(* Logix 5000 project; controller PLC_MCC1300_75F1 vendor 1 type 14 code 166 rev 32.11; software revision 32.04; part 31 of 83 *)
(* tags used below, declared in another part *)
   B70 : DINT[13];
   BENCH_MASTERUP : ALIAS FOR I[73].6;
   C5 : COUNTER[51];
   I : INT[128];   // Local Input Updates Input Slot 2
   KD_N_MOVIN : ALIAS FOR N14[256].0;
   KD_N_MOVOUT : ALIAS FOR N14[257].0;
   KD_S_MOVIN : ALIAS FOR N14[256].1;
   KD_S_MOVOUT : ALIAS FOR N14[257].1;
   KK_N_MOVDN : ALIAS FOR N14[253].0;
   KK_N_MOVIN : ALIAS FOR N14[254].0;
   KK_N_MOVOUT : ALIAS FOR N14[255].0;
   KK_N_MOVUP : ALIAS FOR N14[252].0;
   KK_S_MOVDN : ALIAS FOR N14[253].1;
   KK_S_MOVIN : ALIAS FOR N14[254].1;
   KK_S_MOVOUT : ALIAS FOR N14[255].1;
   KK_S_MOVUP : ALIAS FOR N14[252].1;
   KNRL_N_AUTO : ALIAS FOR N14[250].0;
   KNRL_N_MANL : ALIAS FOR N14[251].0;
   KNRL_S_AUTO : ALIAS FOR N14[250].1;
   KNRL_S_MANL : ALIAS FOR N14[251].1;
   N11 : DINT[500];
   N12 : DINT[500];
   N14 : DINT[500];
   N214_1 : ALIAS FOR N214[1];
   N26 : DINT[150];
   O : INT[128];
   T4 : TIMER[51];
   TD1_N_MOVIN : ALIAS FOR N14[256].2;
   TD1_N_MOVOUT : ALIAS FOR N14[257].2;
   TD1_S_MOVIN : ALIAS FOR N14[256].3;
   TD1_S_MOVOUT : ALIAS FOR N14[257].3;
   TD2_N_MOVIN : ALIAS FOR N14[256].4;
   TD2_N_MOVOUT : ALIAS FOR N14[257].4;
   TK1_N_MOVDN : ALIAS FOR N14[253].2;
   TK1_N_MOVIN : ALIAS FOR N14[254].2;
   TK1_N_MOVOUT : ALIAS FOR N14[255].2;
   TK1_N_MOVUP : ALIAS FOR N14[252].2;
   TK1_S_MOVDN : ALIAS FOR N14[253].3;
   TK1_S_MOVIN : ALIAS FOR N14[254].3;
   TK1_S_MOVOUT : ALIAS FOR N14[255].3;
   TK1_S_MOVUP : ALIAS FOR N14[252].3;
   TK2_N_MOVDN : ALIAS FOR N14[253].4;
   TK2_N_MOVIN : ALIAS FOR N14[254].4;
   TK2_N_MOVOUT : ALIAS FOR N14[255].4;
   TK2_N_MOVUP : ALIAS FOR N14[252].4;
   TK2_S_MOVDN : ALIAS FOR N14[253].5;
   TK2_S_MOVIN : ALIAS FOR N14[254].5;
   TK2_S_MOVOUT : ALIAS FOR N14[255].5;
   TK2_S_MOVUP : ALIAS FOR N14[252].5;
   TMP_d : DINT;
   TZ1_N_AUTO : ALIAS FOR N14[250].2;
   TZ1_N_MANL : ALIAS FOR N14[251].2;
   TZ1_S_AUTO : ALIAS FOR N14[250].3;
   TZ1_S_MANL : ALIAS FOR N14[251].3;
   TZ2_N_AUTO : ALIAS FOR N14[250].4;
   TZ2_N_MANL : ALIAS FOR N14[251].4;
   TZ2_S_AUTO : ALIAS FOR N14[250].5;
   TZ2_S_MANL : ALIAS FOR N14[251].5;
   VIS_OUTPT_OFF : ALIAS FOR N27[60].2;
   VIS_SYS_STOPPED : ALIAS FOR N27[60].1;
(* MainProgram, continued *)

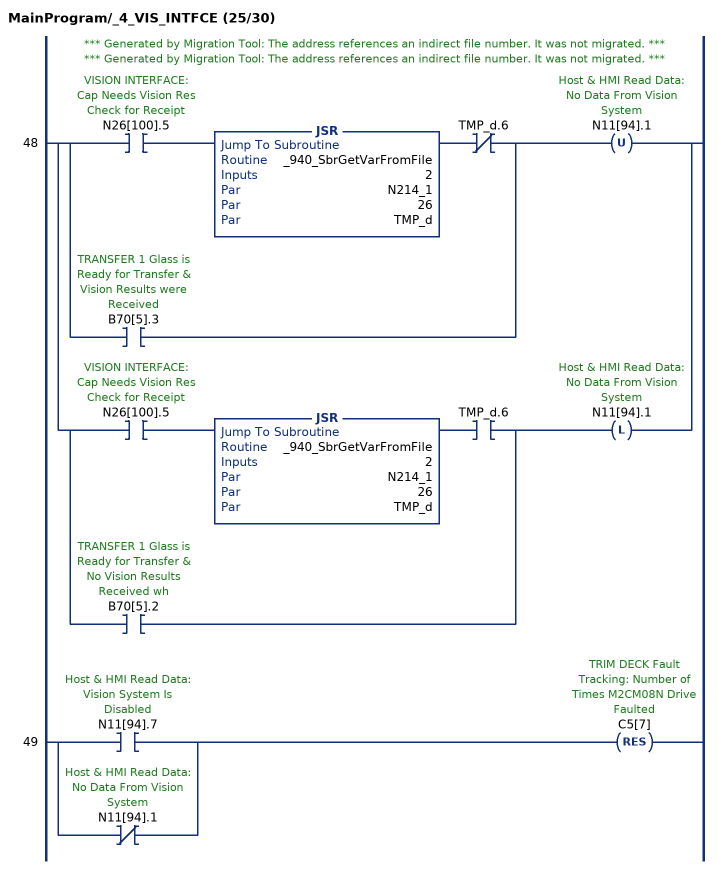
   [picture p426: MainProgram/_4_VIS_INTFCE rungs 48-49]
   // *** Generated by Migration Tool: The address references an indirect file number. It was not migrated. ***
   // *** Generated by Migration Tool: The address references an indirect file number. It was not migrated. ***
   48: [[XIC(N26[100].5) JSR(_940_SbrGetVarFromFile,2,N214_1,26,TMP_d) XIO(TMP_d.6) ,XIC(B70[5].3) ] OTU(N11[94].1) ,[XIC(N26[100].5) JSR(_940_SbrGetVarFromFile,2,N214_1,26,TMP_d) XIC(TMP_d.6) ,XIC(B70[5].2) ] OTL(N11[94].1) ];
   49: [XIC(N11[94].7) ,XIO(N11[94].1) ]RES(C5[7]);
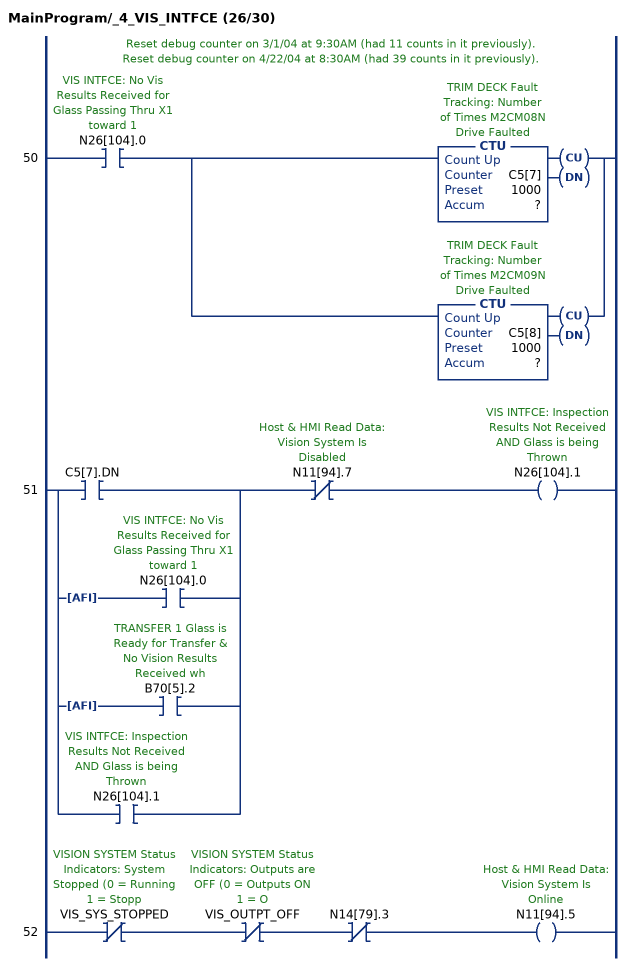
   // Reset debug counter on 3/1/04 at 9:30AM (had 11 counts in it previously).
   // Reset debug counter on 4/22/04 at 8:30AM (had 39 counts in it previously).
   50: XIC(N26[104].0)[CTU(C5[7],?,?) ,CTU(C5[8],?,?) ];
   51: [XIC(C5[7].DN) ,AFI() XIC(N26[104].0) ,AFI() XIC(B70[5].2) ,XIC(N26[104].1) ]XIO(N11[94].7)OTE(N26[104].1);
   52: XIO(VIS_SYS_STOPPED)XIO(VIS_OUTPT_OFF)XIO(N14[79].3)OTE(N11[94].5);
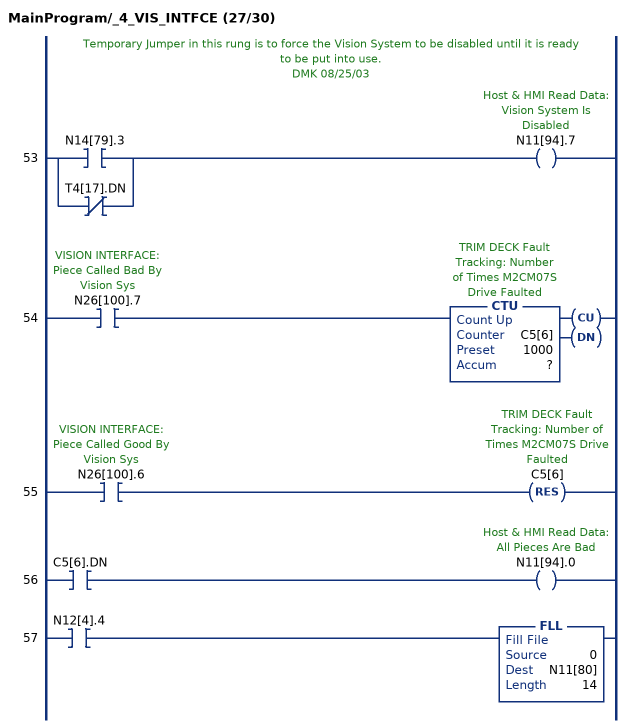
   // Temporary Jumper in this rung is to force the Vision System to be disabled until it is ready to be put into use.
   // DMK 08/25/03
   53: [XIC(N14[79].3) ,XIO(T4[17].DN) ]OTE(N11[94].7);
   54: XIC(N26[100].7)CTU(C5[6],?,?);
   55: XIC(N26[100].6)RES(C5[6]);
   56: XIC(C5[6].DN)OTE(N11[94].0);
   57: XIC(N12[4].4)FLL(0,N11[80],14);
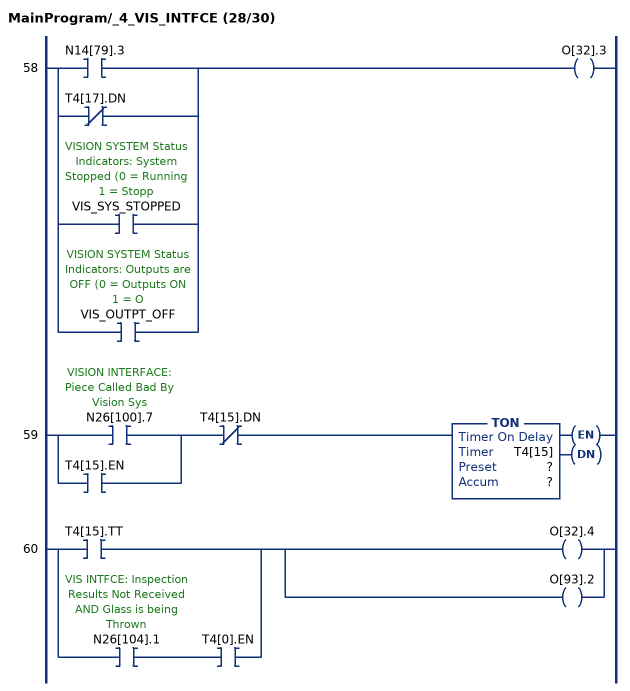
   58: [XIC(N14[79].3) ,XIO(T4[17].DN) ,XIC(VIS_SYS_STOPPED) ,XIC(VIS_OUTPT_OFF) ]OTE(O[32].3);
   59: [XIC(N26[100].7) ,XIC(T4[15].EN) ]XIO(T4[15].DN)TON(T4[15],?,?);
   60: [XIC(T4[15].TT) ,XIC(N26[104].1) XIC(T4[0].EN) ][OTE(O[32].4) ,OTE(O[93].2) ];
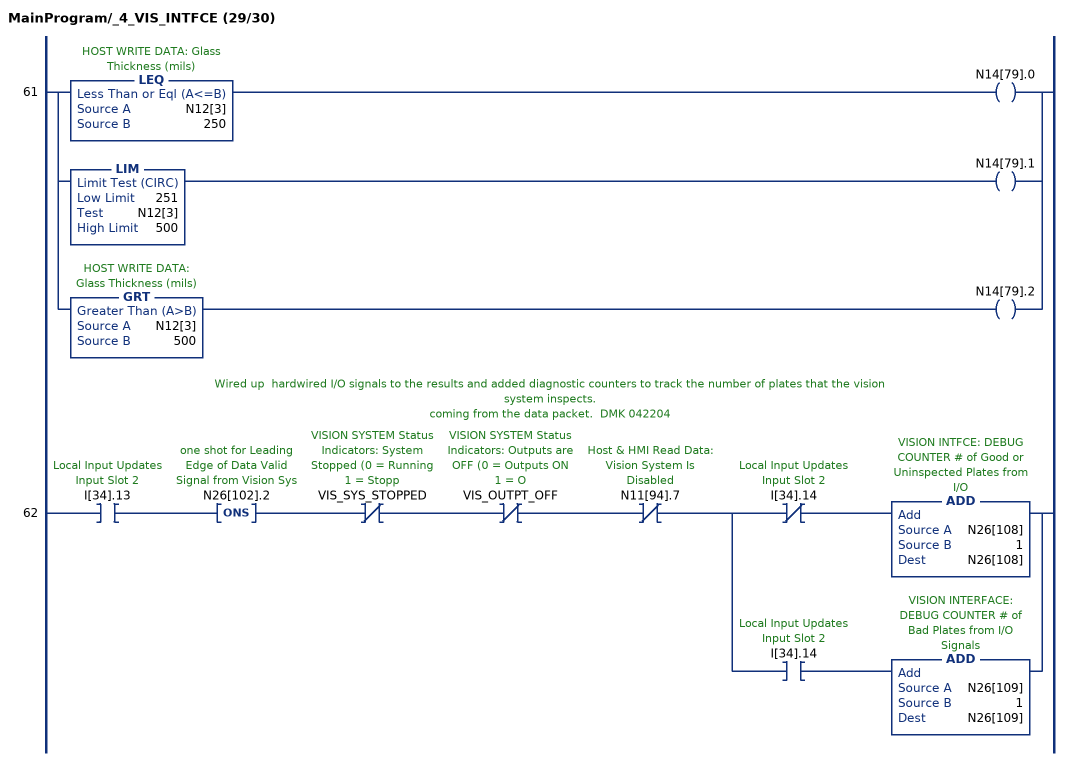
   61: [LEQ(N12[3],250) OTE(N14[79].0) ,LIM(251,N12[3],500) OTE(N14[79].1) ,GRT(N12[3],500) OTE(N14[79].2) ];
   // Wired up  hardwired I/O signals to the results and added diagnostic counters to track the number of plates that the vision
   // system inspects.
   // coming from the data packet.  DMK 042204
   62: XIC(I[34].13)ONS(N26[102].2)XIO(VIS_SYS_STOPPED)XIO(VIS_OUTPT_OFF)XIO(N11[94].7)[XIO(I[34].14) ADD(N26[108],1,N26[108]) ,XIC(I[34].14) ADD(N26[109],1,N26[109]) ];
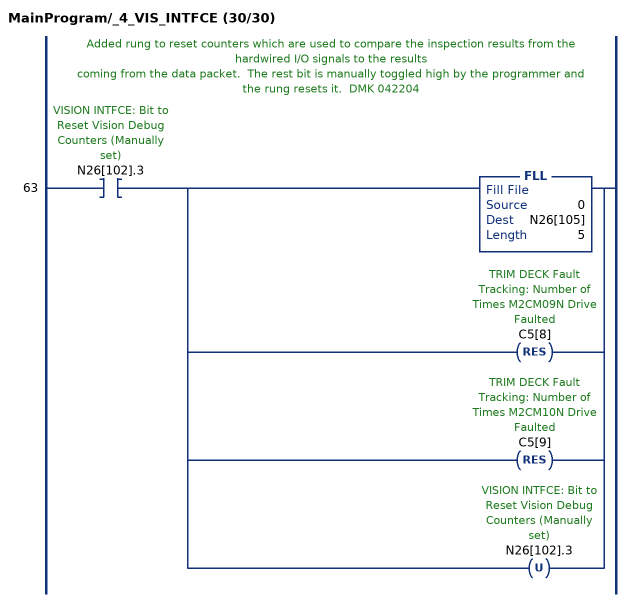
   // Added rung to reset counters which are used to compare the inspection results from the hardwired I/O signals to the results
   // coming from the data packet.  The rest bit is manually toggled high by the programmer and the rung resets it.  DMK 042204
   63: XIC(N26[102].3)[FLL(0,N26[105],5) ,RES(C5[8]) ,RES(C5[9]) ,OTU(N26[102].3) ];
END_ROUTINE

ROUTINE _70_LADDER   (* ladder *)
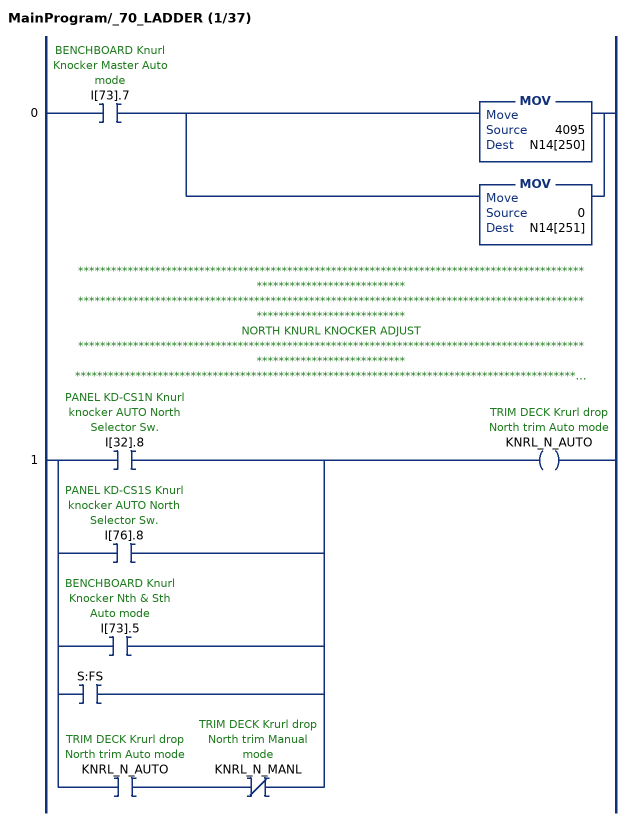
   0: XIC(I[73].7)[MOV(4095,N14[250]) ,MOV(0,N14[251]) ];
   // ***********************************************************************************************************************
   // ***********************************************************************************************************************
   //                                              NORTH KNURL KNOCKER ADJUST
   // ***********************************************************************************************************************
   // ***********************************************************************************************************************
   // North knurl knocker auto mode select
   1: [[XIC(I[32].8) ,XIC(I[76].8) ,XIC(I[73].5) ,XIC(S:FS) ] ,XIC(KNRL_N_AUTO) XIO(KNRL_N_MANL) ]OTE(KNRL_N_AUTO);
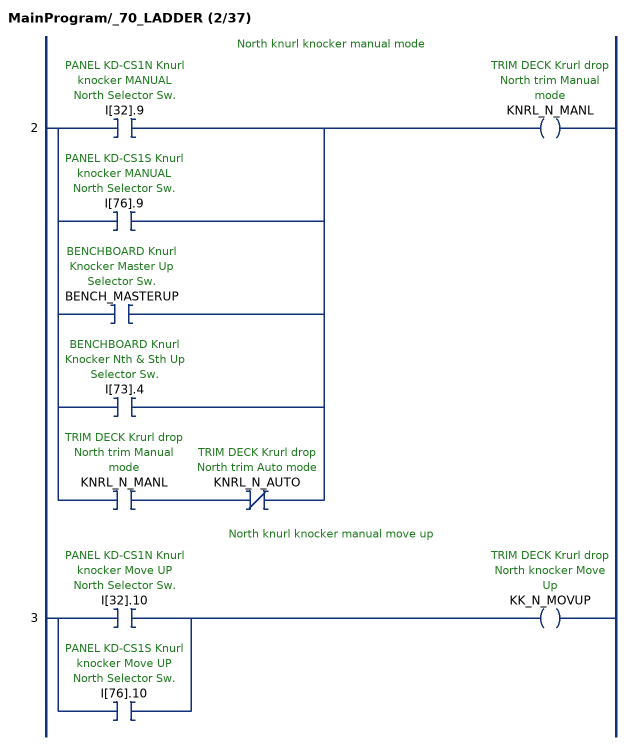
   // North knurl knocker manual mode
   2: [[XIC(I[32].9) ,XIC(I[76].9) ,XIC(BENCH_MASTERUP) ,XIC(I[73].4) ] ,XIC(KNRL_N_MANL) XIO(KNRL_N_AUTO) ]OTE(KNRL_N_MANL);
   // North knurl knocker manual move up
   3: [XIC(I[32].10) ,XIC(I[76].10) ]OTE(KK_N_MOVUP);
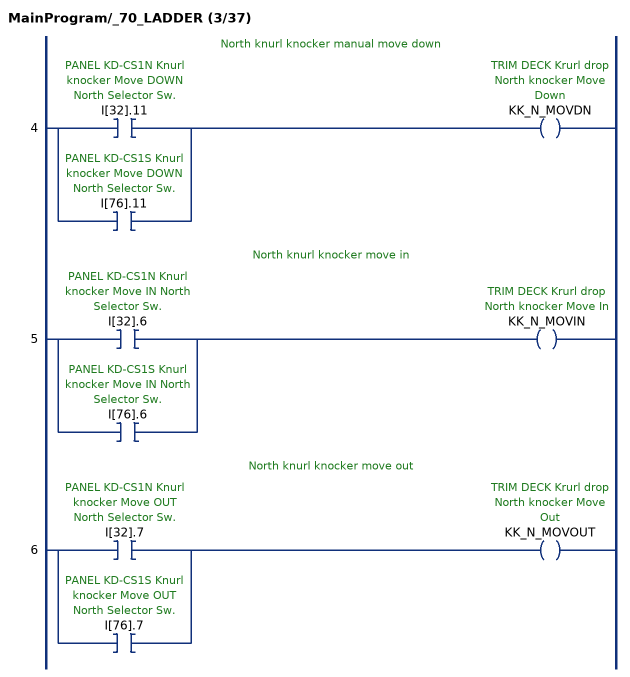
   // North knurl knocker manual move down
   4: [XIC(I[32].11) ,XIC(I[76].11) ]OTE(KK_N_MOVDN);
   // North knurl knocker move in
   5: [XIC(I[32].6) ,XIC(I[76].6) ]OTE(KK_N_MOVIN);
   // North knurl knocker move out
   6: [XIC(I[32].7) ,XIC(I[76].7) ]OTE(KK_N_MOVOUT);
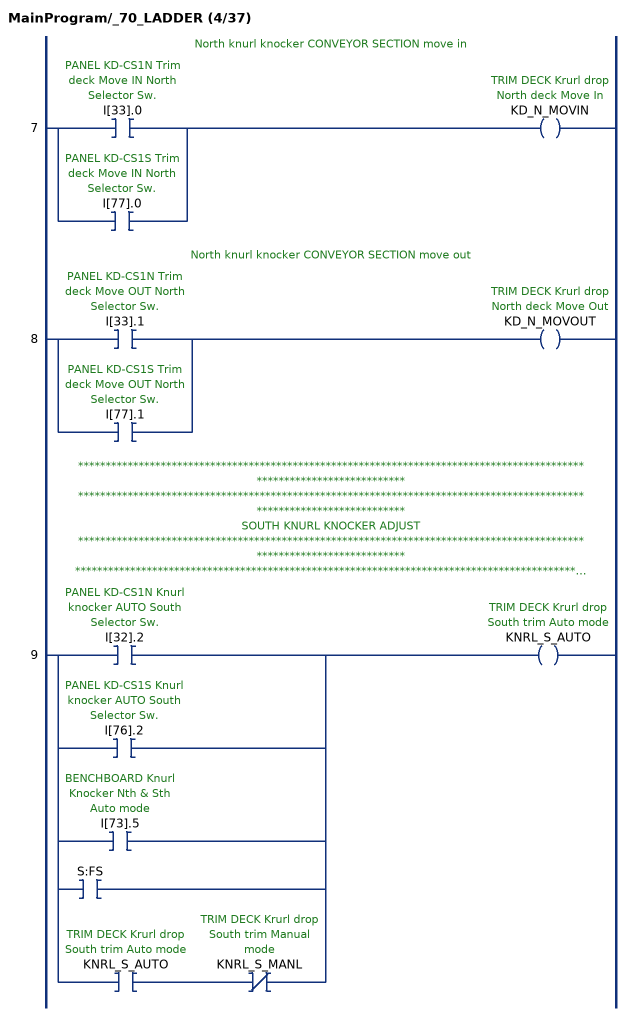
   // North knurl knocker CONVEYOR SECTION move in
   7: [XIC(I[33].0) ,XIC(I[77].0) ]OTE(KD_N_MOVIN);
   // North knurl knocker CONVEYOR SECTION move out
   8: [XIC(I[33].1) ,XIC(I[77].1) ]OTE(KD_N_MOVOUT);
   // ***********************************************************************************************************************
   // ***********************************************************************************************************************
   //                                              SOUTH KNURL KNOCKER ADJUST
   // ***********************************************************************************************************************
   // ***********************************************************************************************************************
   // South knurl knocker auto mode
   9: [[XIC(I[32].2) ,XIC(I[76].2) ,XIC(I[73].5) ,XIC(S:FS) ] ,XIC(KNRL_S_AUTO) XIO(KNRL_S_MANL) ]OTE(KNRL_S_AUTO);
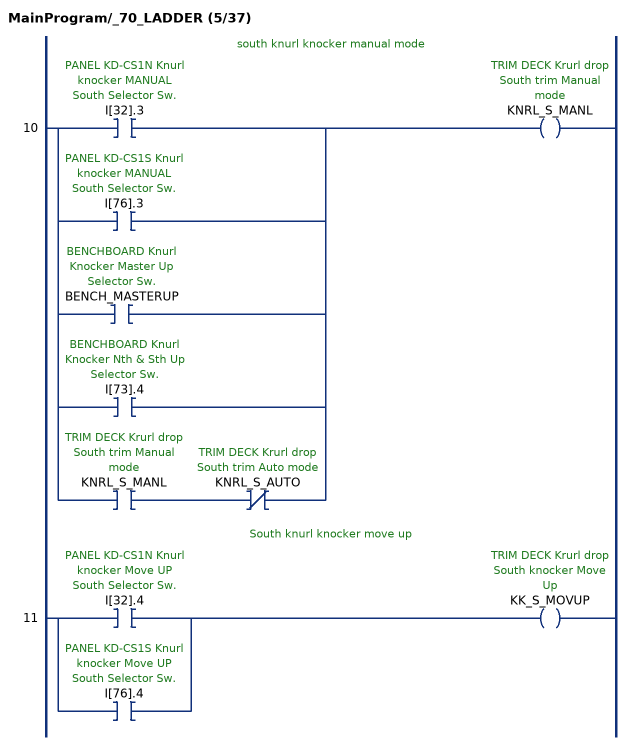
   // south knurl knocker manual mode
   10: [[XIC(I[32].3) ,XIC(I[76].3) ,XIC(BENCH_MASTERUP) ,XIC(I[73].4) ] ,XIC(KNRL_S_MANL) XIO(KNRL_S_AUTO) ]OTE(KNRL_S_MANL);
   // South knurl knocker move up
   11: [XIC(I[32].4) ,XIC(I[76].4) ]OTE(KK_S_MOVUP);
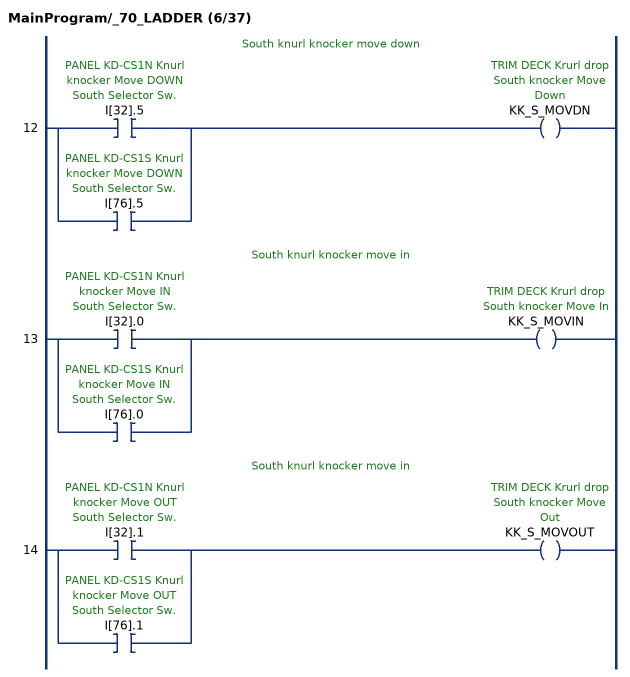
   // South knurl knocker move down
   12: [XIC(I[32].5) ,XIC(I[76].5) ]OTE(KK_S_MOVDN);
   // South knurl knocker move in
   13: [XIC(I[32].0) ,XIC(I[76].0) ]OTE(KK_S_MOVIN);
   // South knurl knocker move in
   14: [XIC(I[32].1) ,XIC(I[76].1) ]OTE(KK_S_MOVOUT);
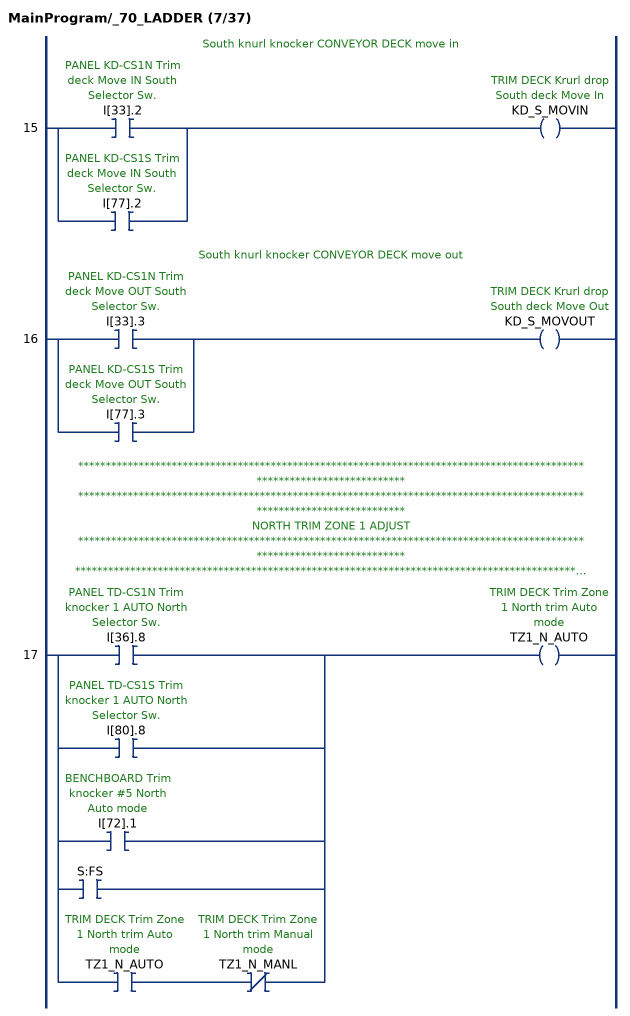
   // South knurl knocker CONVEYOR DECK move in
   15: [XIC(I[33].2) ,XIC(I[77].2) ]OTE(KD_S_MOVIN);
   // South knurl knocker CONVEYOR DECK move out
   16: [XIC(I[33].3) ,XIC(I[77].3) ]OTE(KD_S_MOVOUT);
   // ***********************************************************************************************************************
   // ***********************************************************************************************************************
   //                                              NORTH TRIM ZONE 1 ADJUST
   // ***********************************************************************************************************************
   // ***********************************************************************************************************************
   // North trim knocker 1 auto mode
   17: [[XIC(I[36].8) ,XIC(I[80].8) ,XIC(I[72].1) ,XIC(S:FS) ] ,XIC(TZ1_N_AUTO) XIO(TZ1_N_MANL) ]OTE(TZ1_N_AUTO);
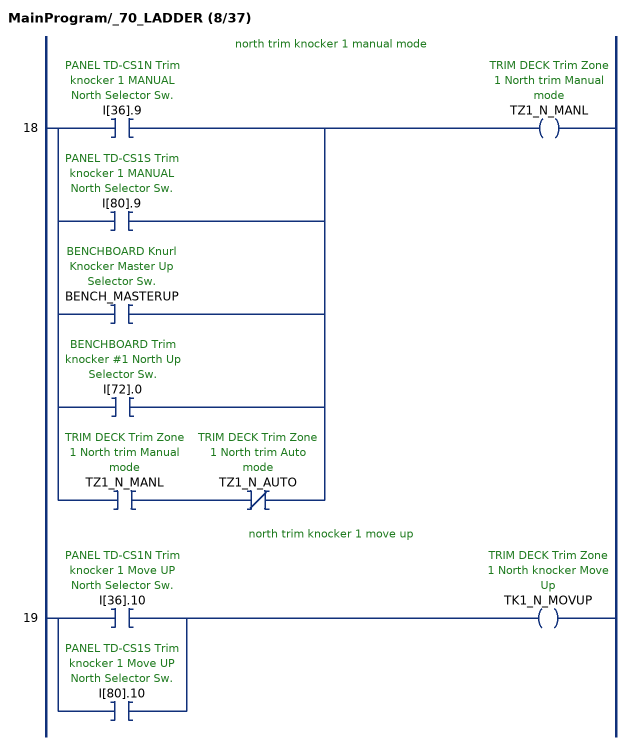
   // north trim knocker 1 manual mode
   18: [[XIC(I[36].9) ,XIC(I[80].9) ,XIC(BENCH_MASTERUP) ,XIC(I[72].0) ] ,XIC(TZ1_N_MANL) XIO(TZ1_N_AUTO) ]OTE(TZ1_N_MANL);
   // north trim knocker 1 move up
   19: [XIC(I[36].10) ,XIC(I[80].10) ]OTE(TK1_N_MOVUP);
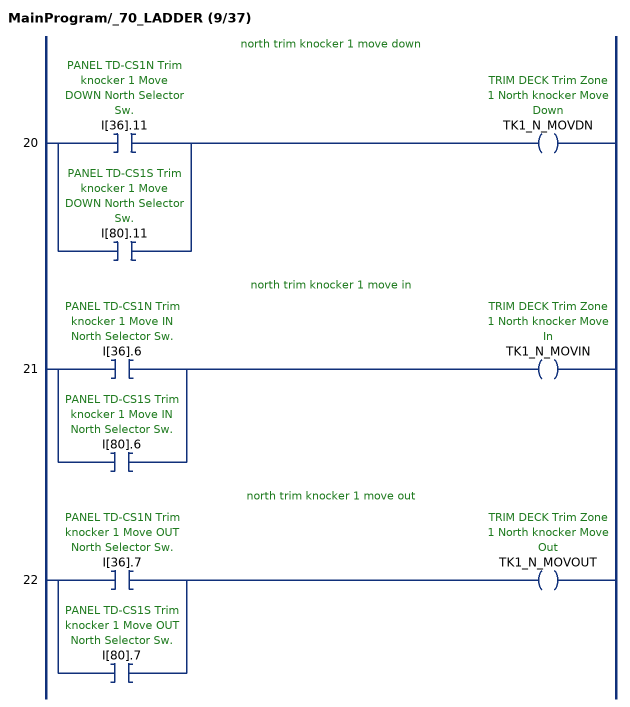
   // north trim knocker 1 move down
   20: [XIC(I[36].11) ,XIC(I[80].11) ]OTE(TK1_N_MOVDN);
   // north trim knocker 1 move in
   21: [XIC(I[36].6) ,XIC(I[80].6) ]OTE(TK1_N_MOVIN);
   // north trim knocker 1 move out
   22: [XIC(I[36].7) ,XIC(I[80].7) ]OTE(TK1_N_MOVOUT);
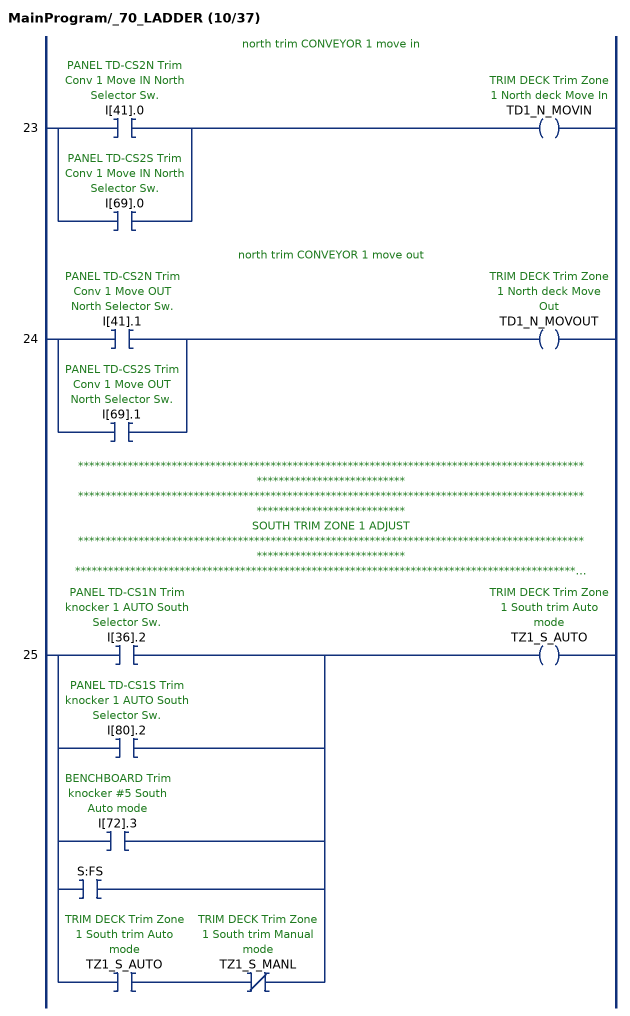
   // north trim CONVEYOR 1 move in
   23: [XIC(I[41].0) ,XIC(I[69].0) ]OTE(TD1_N_MOVIN);
   // north trim CONVEYOR 1 move out
   24: [XIC(I[41].1) ,XIC(I[69].1) ]OTE(TD1_N_MOVOUT);
   // ***********************************************************************************************************************
   // ***********************************************************************************************************************
   //                                              SOUTH TRIM ZONE 1 ADJUST
   // ***********************************************************************************************************************
   // ***********************************************************************************************************************
   // South trim knocker 1 auto mode
   25: [[XIC(I[36].2) ,XIC(I[80].2) ,XIC(I[72].3) ,XIC(S:FS) ] ,XIC(TZ1_S_AUTO) XIO(TZ1_S_MANL) ]OTE(TZ1_S_AUTO);
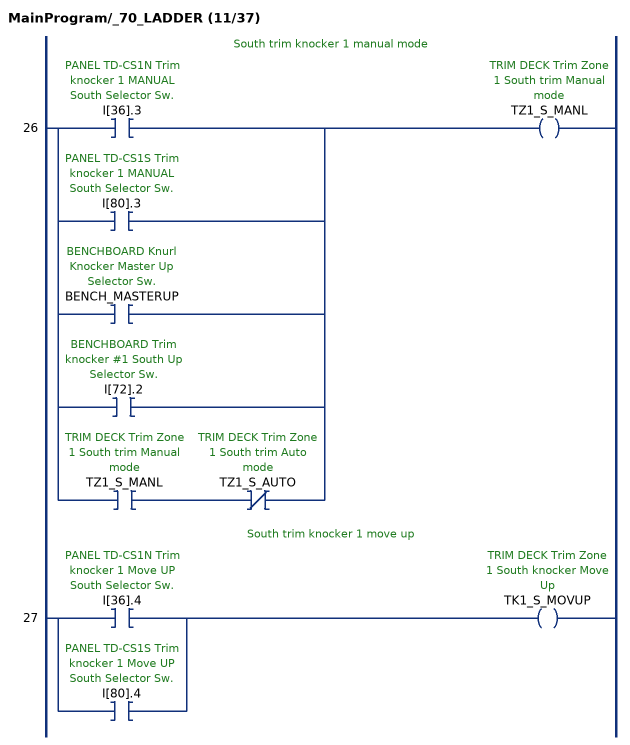
   // South trim knocker 1 manual mode
   26: [[XIC(I[36].3) ,XIC(I[80].3) ,XIC(BENCH_MASTERUP) ,XIC(I[72].2) ] ,XIC(TZ1_S_MANL) XIO(TZ1_S_AUTO) ]OTE(TZ1_S_MANL);
   // South trim knocker 1 move up
   27: [XIC(I[36].4) ,XIC(I[80].4) ]OTE(TK1_S_MOVUP);
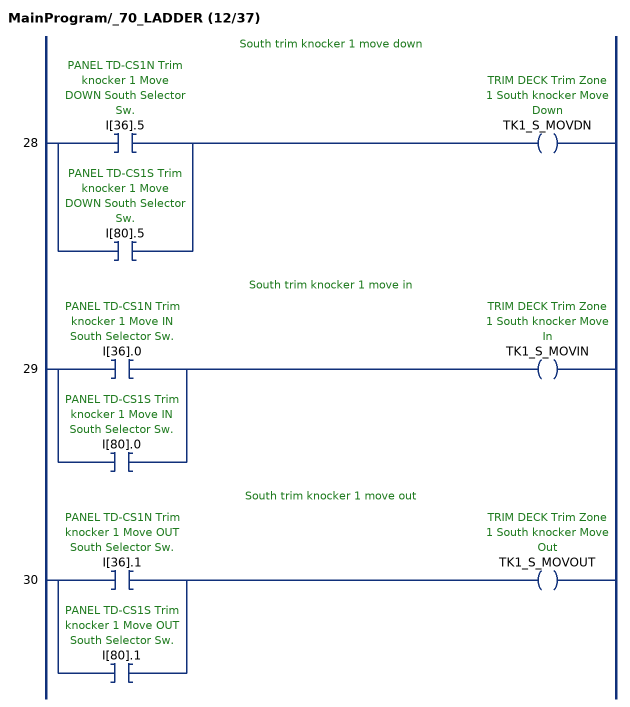
   // South trim knocker 1 move down
   28: [XIC(I[36].5) ,XIC(I[80].5) ]OTE(TK1_S_MOVDN);
   // South trim knocker 1 move in
   29: [XIC(I[36].0) ,XIC(I[80].0) ]OTE(TK1_S_MOVIN);
   // South trim knocker 1 move out
   30: [XIC(I[36].1) ,XIC(I[80].1) ]OTE(TK1_S_MOVOUT);
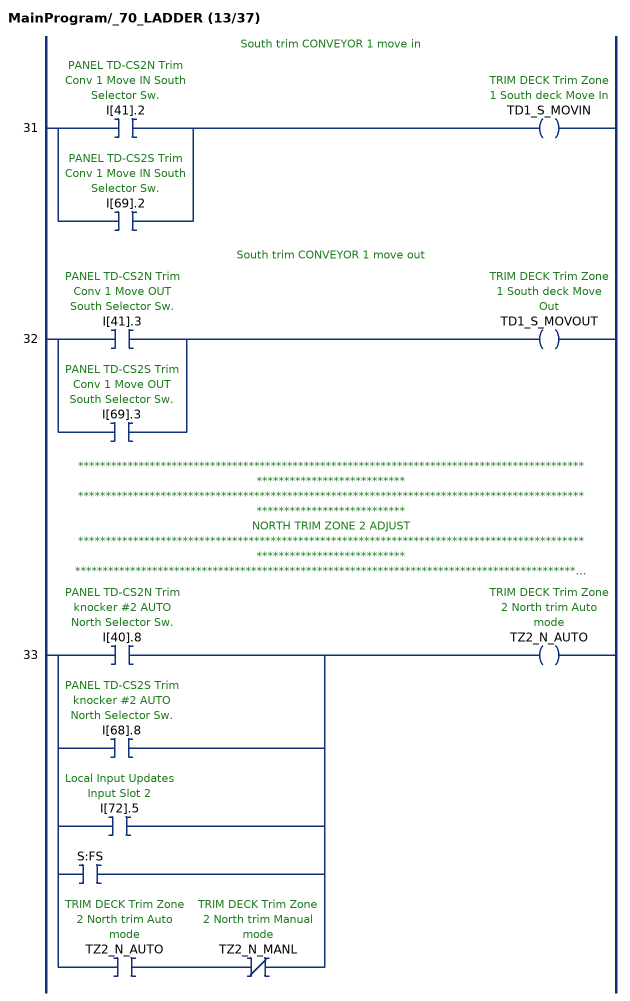
   // South trim CONVEYOR 1 move in
   31: [XIC(I[41].2) ,XIC(I[69].2) ]OTE(TD1_S_MOVIN);
   // South trim CONVEYOR 1 move out
   32: [XIC(I[41].3) ,XIC(I[69].3) ]OTE(TD1_S_MOVOUT);
   // ***********************************************************************************************************************
   // ***********************************************************************************************************************
   //                                              NORTH TRIM ZONE 2 ADJUST
   // ***********************************************************************************************************************
   // ***********************************************************************************************************************
   // North trim knocker 2 auto mode
   33: [[XIC(I[40].8) ,XIC(I[68].8) ,XIC(I[72].5) ,XIC(S:FS) ] ,XIC(TZ2_N_AUTO) XIO(TZ2_N_MANL) ]OTE(TZ2_N_AUTO);
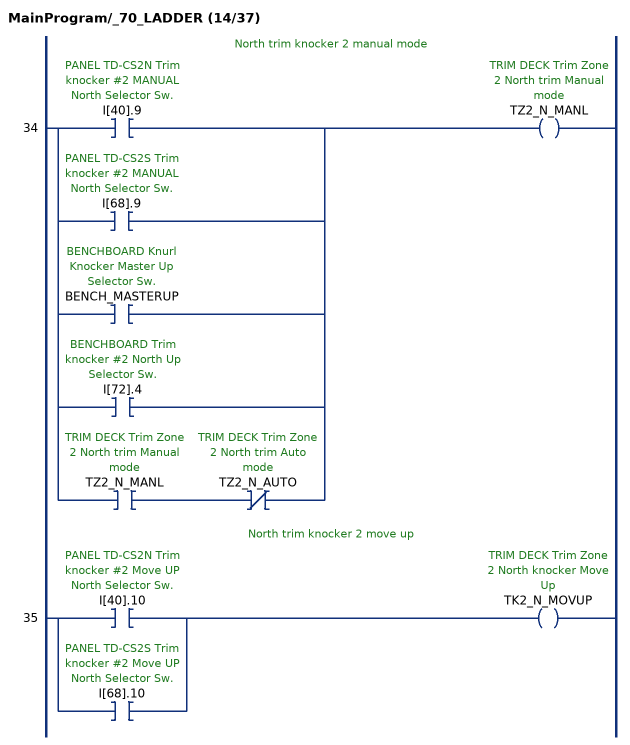
   // North trim knocker 2 manual mode
   34: [[XIC(I[40].9) ,XIC(I[68].9) ,XIC(BENCH_MASTERUP) ,XIC(I[72].4) ] ,XIC(TZ2_N_MANL) XIO(TZ2_N_AUTO) ]OTE(TZ2_N_MANL);
   // North trim knocker 2 move up
   35: [XIC(I[40].10) ,XIC(I[68].10) ]OTE(TK2_N_MOVUP);
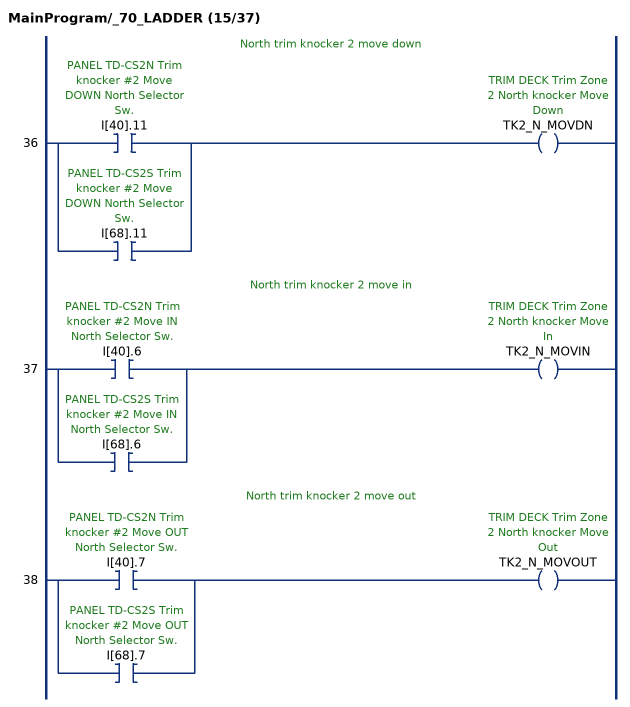
   // North trim knocker 2 move down
   36: [XIC(I[40].11) ,XIC(I[68].11) ]OTE(TK2_N_MOVDN);
   // North trim knocker 2 move in
   37: [XIC(I[40].6) ,XIC(I[68].6) ]OTE(TK2_N_MOVIN);
   // North trim knocker 2 move out
   38: [XIC(I[40].7) ,XIC(I[68].7) ]OTE(TK2_N_MOVOUT);
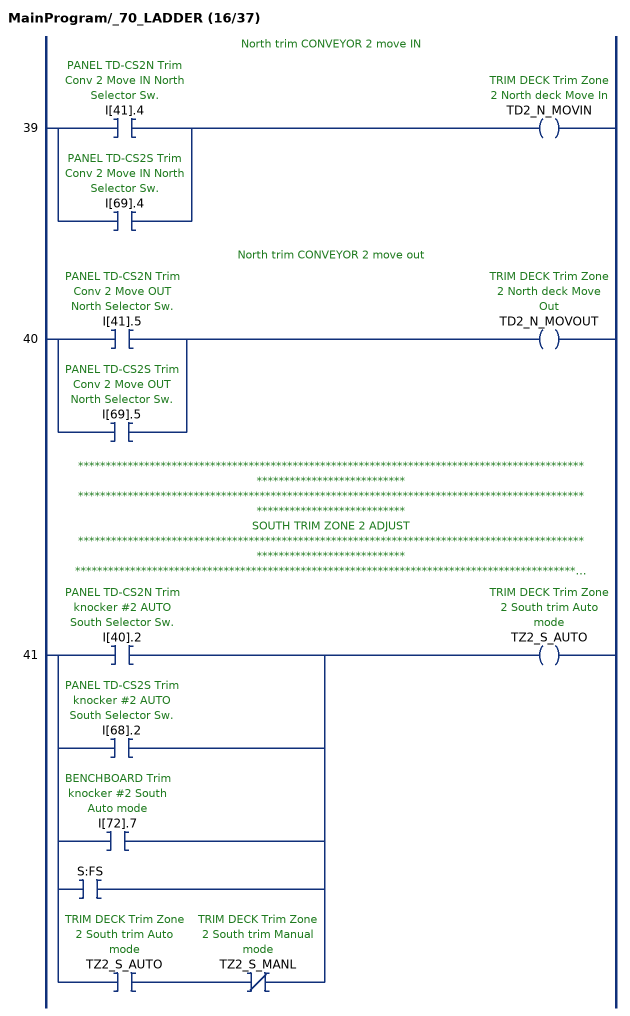
   // North trim CONVEYOR 2 move IN
   39: [XIC(I[41].4) ,XIC(I[69].4) ]OTE(TD2_N_MOVIN);
   // North trim CONVEYOR 2 move out
   40: [XIC(I[41].5) ,XIC(I[69].5) ]OTE(TD2_N_MOVOUT);
   // ***********************************************************************************************************************
   // ***********************************************************************************************************************
   //                                              SOUTH TRIM ZONE 2 ADJUST
   // ***********************************************************************************************************************
   // ***********************************************************************************************************************
   // South trim knocker 2 auto mode
   41: [[XIC(I[40].2) ,XIC(I[68].2) ,XIC(I[72].7) ,XIC(S:FS) ] ,XIC(TZ2_S_AUTO) XIO(TZ2_S_MANL) ]OTE(TZ2_S_AUTO);
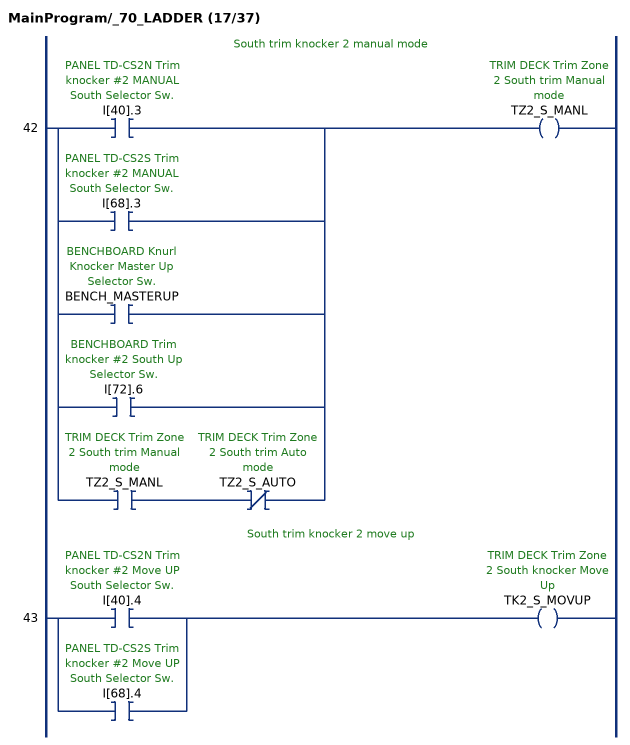
   // South trim knocker 2 manual mode
   42: [[XIC(I[40].3) ,XIC(I[68].3) ,XIC(BENCH_MASTERUP) ,XIC(I[72].6) ] ,XIC(TZ2_S_MANL) XIO(TZ2_S_AUTO) ]OTE(TZ2_S_MANL);
   // South trim knocker 2 move up
   43: [XIC(I[40].4) ,XIC(I[68].4) ]OTE(TK2_S_MOVUP);
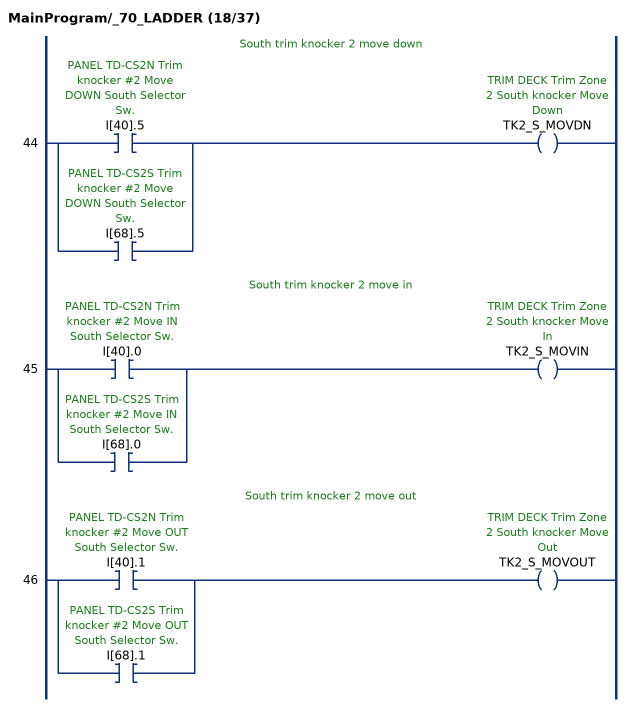
   // South trim knocker 2 move down
   44: [XIC(I[40].5) ,XIC(I[68].5) ]OTE(TK2_S_MOVDN);
   // South trim knocker 2 move in
   45: [XIC(I[40].0) ,XIC(I[68].0) ]OTE(TK2_S_MOVIN);
   // South trim knocker 2 move out
   46: [XIC(I[40].1) ,XIC(I[68].1) ]OTE(TK2_S_MOVOUT);
